TYPE "KP8 Driver: Parameters: 1 Button"
   STRUCT
      activate : Bool;   // true = button on, flase = button off
      cOn1 : String[10];   // color when button is in pressed state. valid entries: 'red', 'green', 'blue', 'yellow', 'white', 'off'
      cOn2 : String[10];   // second flash color when button is pressed and flashing is enabled. valid entries: 'red', 'green', 'blue', 'yellow', 'white', 'off'
      cOff : String[10];   // color when button is in un-pressed state. valid entries: 'red', 'green', 'blue', 'yellow', 'white', 'off'
      flash : Bool;   // false = color 1, true = color 2. set to clock bit to flash at that rate
      group : Int;   // 0 disables. buttons in groups have a mutually exclusive 'on' state.
      mode : Bool;   // true = maintained, fales = momentary
   END_STRUCT;
END_TYPE

TYPE "Selectable Wips"
   STRUCT
      count : Int;
      wips : Array[0.."wipCount"] of DInt;
   END_STRUCT;
END_TYPE

TYPE "Recipe: PN Text Library"
VERSION : 0.1
   STRUCT
      pnText : Array[0.."pnLibCount"] of WString["sStringLen"];
   END_STRUCT;
END_TYPE

TYPE "Selected Wips"
   STRUCT
      count : Int;
      wips : Array[0.."wipCount"] of DInt;
   END_STRUCT;
END_TYPE

TYPE "Selected Buttons"
   STRUCT
      btns : Array[0.."btnCount"] of Bool;
      count : Int;
   END_STRUCT;
END_TYPE

TYPE "KP8 Driver: Button States"
   STRUCT
      btn : Array[0..7] of Bool;
   END_STRUCT;
END_TYPE

TYPE "KP8 Driver: Parameters: 8 Buttons"
   STRUCT
      btn : Array[0..7] of "KP8 Driver: Parameters: 1 Button";
   END_STRUCT;
END_TYPE

TYPE "KP8 Driver: Feedback Data"
   STRUCT
      acutal : "KP8 Driver: Button States";
      falling : "KP8 Driver: Button States";
      rising : "KP8 Driver: Button States";
   END_STRUCT;
END_TYPE

TYPE "Setting Meta Data"
   STRUCT
      selectable_stations : "Selectable Stations";
      selectable_wips : "Selectable Wips";
      selected_btns : "Selected Buttons";
      selected_stations : "Selected Stations";
      selected_wips : "Selected Wips";
      selection_change : "Station Selection Change";
   END_STRUCT;
END_TYPE

TYPE "Nav Bar Data"
   STRUCT
      hmi : "Nav Bar Data: HMI";
      plc : "Nav Bar Data: PLC";
   END_STRUCT;
END_TYPE

TYPE "Intersecting WIPs Arrays"
   STRUCT
      count : Int;
      WIPS_intersection : Array[0.."wipCount"] of DInt;
   END_STRUCT;
END_TYPE

TYPE "Initialize Excel Data: States"
   STRUCT
      active_wip_to_hmi_station_list : Bool;
      active_wip_to_master_station_list : Bool;
      pn_code_to_kp8_station : Bool;
      pn_code_to_saved_wips : Bool;
      wip_code_to_saved_wips : Bool;
   END_STRUCT;
END_TYPE

DATA_BLOCK "EMP IDB"   // DB1
{ S7_Optimized_Access := 'TRUE' }
VERSION : 0.1
// stored: InstanceOfName EMP
"EMP"
BEGIN
   "inst HMI Station"."inst HMI Station: Wip Selection".rowIndicies[1] := 1;
   "inst HMI Station"."inst HMI Station: Wip Selection".rowIndicies[2] := 2;
   "inst HMI Station"."inst HMI Station: Wip Selection".rowIndicies[3] := 3;
   "inst HMI Station"."inst HMI Station: Wip Selection".rowIndicies[4] := 4;
   "inst HMI Station"."inst HMI Station: Wip Selection".rowIndicies[5] := 5;
END_DATA_BLOCK

DATA_BLOCK "Debug"   // DB7
{ S7_Optimized_Access := 'TRUE' }
VERSION : 0.1
   VAR
      nullCheck : Array[0.."wipCount"] of DInt;
   END_VAR
BEGIN
END_DATA_BLOCK

// folder: From Excel

DATA_BLOCK "From Excel: Codes"   // DB12
{ S7_Optimized_Access := 'TRUE' }
VERSION : 0.1
BEGIN
   kp8Stns[0].pnCode[0] := 0;
   kp8Stns[0].pnCode[1] := 0;
   kp8Stns[0].pnCode[2] := 0;
   kp8Stns[0].pnCode[3] := 172000;
   kp8Stns[0].pnCode[4] := 0;
   kp8Stns[0].pnCode[5] := 0;
   kp8Stns[0].pnCode[6] := 0;
   kp8Stns[0].pnCode[7] := 168000;
   kp8Stns[1].pnCode[0] := 0;
   kp8Stns[1].pnCode[1] := 0;
   kp8Stns[1].pnCode[2] := 183000;
   kp8Stns[1].pnCode[3] := 209000;
   kp8Stns[1].pnCode[4] := 0;
   kp8Stns[1].pnCode[5] := 0;
   kp8Stns[1].pnCode[6] := 180000;
   kp8Stns[1].pnCode[7] := 166000;
   kp8Stns[2].pnCode[0] := 0;
   kp8Stns[2].pnCode[1] := 182000;
   kp8Stns[2].pnCode[2] := 181000;
   kp8Stns[2].pnCode[3] := 215000;
   kp8Stns[2].pnCode[4] := 0;
   kp8Stns[2].pnCode[5] := 184000;
   kp8Stns[2].pnCode[6] := 216000;
   kp8Stns[2].pnCode[7] := 214000;
   kp8Stns[3].pnCode[0] := 0;
   kp8Stns[3].pnCode[1] := 192000;
   kp8Stns[3].pnCode[2] := 191000;
   kp8Stns[3].pnCode[3] := 188000;
   kp8Stns[3].pnCode[4] := 0;
   kp8Stns[3].pnCode[5] := 190000;
   kp8Stns[3].pnCode[6] := 187000;
   kp8Stns[3].pnCode[7] := 189000;
   kp8Stns[4].pnCode[0] := 0;
   kp8Stns[4].pnCode[1] := 0;
   kp8Stns[4].pnCode[2] := 0;
   kp8Stns[4].pnCode[3] := 0;
   kp8Stns[4].pnCode[4] := 0;
   kp8Stns[4].pnCode[5] := 0;
   kp8Stns[4].pnCode[6] := 0;
   kp8Stns[4].pnCode[7] := 194000;
   kp8Stns[5].pnCode[0] := 0;
   kp8Stns[5].pnCode[1] := 193000;
   kp8Stns[5].pnCode[2] := 195000;
   kp8Stns[5].pnCode[3] := 176000;
   kp8Stns[5].pnCode[4] := 0;
   kp8Stns[5].pnCode[5] := 196000;
   kp8Stns[5].pnCode[6] := 177000;
   kp8Stns[5].pnCode[7] := 175000;
   kp8Stns[6].pnCode[0] := 0;
   kp8Stns[6].pnCode[1] := 208000;
   kp8Stns[6].pnCode[2] := 207000;
   kp8Stns[6].pnCode[3] := 210000;
   kp8Stns[6].pnCode[4] := 0;
   kp8Stns[6].pnCode[5] := 211000;
   kp8Stns[6].pnCode[6] := 206000;
   kp8Stns[6].pnCode[7] := 205000;
   kp8Stns[7].pnCode[0] := 0;
   kp8Stns[7].pnCode[1] := 0;
   kp8Stns[7].pnCode[2] := 0;
   kp8Stns[7].pnCode[3] := 174000;
   kp8Stns[7].pnCode[4] := 0;
   kp8Stns[7].pnCode[5] := 0;
   kp8Stns[7].pnCode[6] := 167000;
   kp8Stns[7].pnCode[7] := 169000;
   kp8Stns[8].pnCode[0] := 0;
   kp8Stns[8].pnCode[1] := 0;
   kp8Stns[8].pnCode[2] := 0;
   kp8Stns[8].pnCode[3] := 204000;
   kp8Stns[8].pnCode[4] := 0;
   kp8Stns[8].pnCode[5] := 0;
   kp8Stns[8].pnCode[6] := 173000;
   kp8Stns[8].pnCode[7] := 186000;
   kp8Stns[9].pnCode[0] := 0;
   kp8Stns[9].pnCode[1] := 0;
   kp8Stns[9].pnCode[2] := 0;
   kp8Stns[9].pnCode[3] := 213000;
   kp8Stns[9].pnCode[4] := 0;
   kp8Stns[9].pnCode[5] := 0;
   kp8Stns[9].pnCode[6] := 0;
   kp8Stns[9].pnCode[7] := 212000;
   kp8Stns[10].pnCode[0] := 0;
   kp8Stns[10].pnCode[1] := 0;
   kp8Stns[10].pnCode[2] := 0;
   kp8Stns[10].pnCode[3] := 170000;
   kp8Stns[10].pnCode[4] := 0;
   kp8Stns[10].pnCode[5] := 0;
   kp8Stns[10].pnCode[6] := 242000;
   kp8Stns[10].pnCode[7] := 171000;
   kp8Stns[11].pnCode[0] := 0;
   kp8Stns[11].pnCode[1] := 0;
   kp8Stns[11].pnCode[2] := 0;
   kp8Stns[11].pnCode[3] := 77000;
   kp8Stns[11].pnCode[4] := 0;
   kp8Stns[11].pnCode[5] := 0;
   kp8Stns[11].pnCode[6] := 65000;
   kp8Stns[11].pnCode[7] := 20000;
   kp8Stns[12].pnCode[0] := 0;
   kp8Stns[12].pnCode[1] := 80000;
   kp8Stns[12].pnCode[2] := 86000;
   kp8Stns[12].pnCode[3] := 59000;
   kp8Stns[12].pnCode[4] := 0;
   kp8Stns[12].pnCode[5] := 79000;
   kp8Stns[12].pnCode[6] := 55000;
   kp8Stns[12].pnCode[7] := 54000;
   kp8Stns[13].pnCode[0] := 0;
   kp8Stns[13].pnCode[1] := 0;
   kp8Stns[13].pnCode[2] := 69000;
   kp8Stns[13].pnCode[3] := 89000;
   kp8Stns[13].pnCode[4] := 0;
   kp8Stns[13].pnCode[5] := 0;
   kp8Stns[13].pnCode[6] := 90000;
   kp8Stns[13].pnCode[7] := 88000;
   kp8Stns[14].pnCode[0] := 0;
   kp8Stns[14].pnCode[1] := 0;
   kp8Stns[14].pnCode[2] := 64000;
   kp8Stns[14].pnCode[3] := 87000;
   kp8Stns[14].pnCode[4] := 0;
   kp8Stns[14].pnCode[5] := 63000;
   kp8Stns[14].pnCode[6] := 82000;
   kp8Stns[14].pnCode[7] := 62000;
   kp8Stns[15].pnCode[0] := 0;
   kp8Stns[15].pnCode[1] := 49000;
   kp8Stns[15].pnCode[2] := 76000;
   kp8Stns[15].pnCode[3] := 28000;
   kp8Stns[15].pnCode[4] := 0;
   kp8Stns[15].pnCode[5] := 81000;
   kp8Stns[15].pnCode[6] := 68000;
   kp8Stns[15].pnCode[7] := 74000;
   kp8Stns[16].pnCode[0] := 0;
   kp8Stns[16].pnCode[1] := 0;
   kp8Stns[16].pnCode[2] := 0;
   kp8Stns[16].pnCode[3] := 91000;
   kp8Stns[16].pnCode[4] := 0;
   kp8Stns[16].pnCode[5] := 0;
   kp8Stns[16].pnCode[6] := 93000;
   kp8Stns[16].pnCode[7] := 94067;
   kp8Stns[17].pnCode[0] := 0;
   kp8Stns[17].pnCode[1] := 0;
   kp8Stns[17].pnCode[2] := 83000;
   kp8Stns[17].pnCode[3] := 34000;
   kp8Stns[17].pnCode[4] := 0;
   kp8Stns[17].pnCode[5] := 0;
   kp8Stns[17].pnCode[6] := 75000;
   kp8Stns[17].pnCode[7] := 29000;
   kp8Stns[18].pnCode[0] := 0;
   kp8Stns[18].pnCode[1] := 0;
   kp8Stns[18].pnCode[2] := 0;
   kp8Stns[18].pnCode[3] := 92066;
   kp8Stns[18].pnCode[4] := 0;
   kp8Stns[18].pnCode[5] := 0;
   kp8Stns[18].pnCode[6] := 96026;
   kp8Stns[18].pnCode[7] := 95000;
   kp8Stns[19].pnCode[0] := 0;
   kp8Stns[19].pnCode[1] := 78000;
   kp8Stns[19].pnCode[2] := 85000;
   kp8Stns[19].pnCode[3] := 21000;
   kp8Stns[19].pnCode[4] := 0;
   kp8Stns[19].pnCode[5] := 97000;
   kp8Stns[19].pnCode[6] := 60000;
   kp8Stns[19].pnCode[7] := 48000;
   kp8Stns[20].pnCode[0] := 0;
   kp8Stns[20].pnCode[1] := 0;
   kp8Stns[20].pnCode[2] := 0;
   kp8Stns[20].pnCode[3] := 0;
   kp8Stns[20].pnCode[4] := 0;
   kp8Stns[20].pnCode[5] := 0;
   kp8Stns[20].pnCode[6] := 0;
   kp8Stns[20].pnCode[7] := 244000;
   kp8Stns[21].pnCode[0] := 0;
   kp8Stns[21].pnCode[1] := 0;
   kp8Stns[21].pnCode[2] := 0;
   kp8Stns[21].pnCode[3] := 245000;
   kp8Stns[21].pnCode[4] := 0;
   kp8Stns[21].pnCode[5] := 0;
   kp8Stns[21].pnCode[6] := 0;
   kp8Stns[21].pnCode[7] := 11000;
   kp8Stns[22].pnCode[0] := 0;
   kp8Stns[22].pnCode[1] := 0;
   kp8Stns[22].pnCode[2] := 0;
   kp8Stns[22].pnCode[3] := 22000;
   kp8Stns[22].pnCode[4] := 0;
   kp8Stns[22].pnCode[5] := 0;
   kp8Stns[22].pnCode[6] := 46000;
   kp8Stns[22].pnCode[7] := 61000;
   kp8Stns[23].pnCode[0] := 0;
   kp8Stns[23].pnCode[1] := 0;
   kp8Stns[23].pnCode[2] := 0;
   kp8Stns[23].pnCode[3] := 0;
   kp8Stns[23].pnCode[4] := 0;
   kp8Stns[23].pnCode[5] := 0;
   kp8Stns[23].pnCode[6] := 0;
   kp8Stns[23].pnCode[7] := 12000;
   kp8Stns[24].pnCode[0] := 0;
   kp8Stns[24].pnCode[1] := 0;
   kp8Stns[24].pnCode[2] := 0;
   kp8Stns[24].pnCode[3] := 0;
   kp8Stns[24].pnCode[4] := 0;
   kp8Stns[24].pnCode[5] := 0;
   kp8Stns[24].pnCode[6] := 0;
   kp8Stns[24].pnCode[7] := 27000;
   kp8Stns[25].pnCode[0] := 0;
   kp8Stns[25].pnCode[1] := 0;
   kp8Stns[25].pnCode[2] := 0;
   kp8Stns[25].pnCode[3] := 0;
   kp8Stns[25].pnCode[4] := 0;
   kp8Stns[25].pnCode[5] := 0;
   kp8Stns[25].pnCode[6] := 0;
   kp8Stns[25].pnCode[7] := 56000;
   hmiStns[0].wip[0].wipCode := 6027;
   hmiStns[0].wip[0].pnCode[0] := 0;
   hmiStns[0].wip[0].pnCode[1] := 243000;
   hmiStns[0].wip[0].pnCode[2] := 19000;
   hmiStns[0].wip[0].pnCode[3] := 0;
   hmiStns[0].wip[0].pnCode[4] := 0;
   hmiStns[0].wip[0].pnCode[5] := 0;
   hmiStns[0].wip[0].pnCode[6] := 25000;
   hmiStns[0].wip[0].pnCode[7] := 18000;
   hmiStns[0].wip[1].wipCode := 9007;
   hmiStns[0].wip[1].pnCode[0] := 0;
   hmiStns[0].wip[1].pnCode[1] := 243000;
   hmiStns[0].wip[1].pnCode[2] := 37000;
   hmiStns[0].wip[1].pnCode[3] := 0;
   hmiStns[0].wip[1].pnCode[4] := 0;
   hmiStns[0].wip[1].pnCode[5] := 0;
   hmiStns[0].wip[1].pnCode[6] := 35000;
   hmiStns[0].wip[1].pnCode[7] := 36000;
   hmiStns[0].wip[2].wipCode := 10030;
   hmiStns[0].wip[2].pnCode[0] := 0;
   hmiStns[0].wip[2].pnCode[1] := 243000;
   hmiStns[0].wip[2].pnCode[2] := 40000;
   hmiStns[0].wip[2].pnCode[3] := 0;
   hmiStns[0].wip[2].pnCode[4] := 0;
   hmiStns[0].wip[2].pnCode[5] := 0;
   hmiStns[0].wip[2].pnCode[6] := 38000;
   hmiStns[0].wip[2].pnCode[7] := 39000;
   hmiStns[0].wip[3].wipCode := 11056;
   hmiStns[0].wip[3].pnCode[0] := 0;
   hmiStns[0].wip[3].pnCode[1] := 243000;
   hmiStns[0].wip[3].pnCode[2] := 47000;
   hmiStns[0].wip[3].pnCode[3] := 13000;
   hmiStns[0].wip[3].pnCode[4] := 0;
   hmiStns[0].wip[3].pnCode[5] := 14000;
   hmiStns[0].wip[3].pnCode[6] := 41000;
   hmiStns[0].wip[3].pnCode[7] := 32000;
   hmiStns[0].wip[4].wipCode := 12008;
   hmiStns[0].wip[4].pnCode[0] := 0;
   hmiStns[0].wip[4].pnCode[1] := 243000;
   hmiStns[0].wip[4].pnCode[2] := 45000;
   hmiStns[0].wip[4].pnCode[3] := 0;
   hmiStns[0].wip[4].pnCode[4] := 0;
   hmiStns[0].wip[4].pnCode[5] := 0;
   hmiStns[0].wip[4].pnCode[6] := 35000;
   hmiStns[0].wip[4].pnCode[7] := 36000;
   hmiStns[0].wip[5].wipCode := 13060;
   hmiStns[0].wip[5].pnCode[0] := 0;
   hmiStns[0].wip[5].pnCode[1] := 243000;
   hmiStns[0].wip[5].pnCode[2] := 37000;
   hmiStns[0].wip[5].pnCode[3] := 0;
   hmiStns[0].wip[5].pnCode[4] := 0;
   hmiStns[0].wip[5].pnCode[5] := 0;
   hmiStns[0].wip[5].pnCode[6] := 42000;
   hmiStns[0].wip[5].pnCode[7] := 36000;
   hmiStns[0].wip[6].wipCode := 14061;
   hmiStns[0].wip[6].pnCode[0] := 0;
   hmiStns[0].wip[6].pnCode[1] := 243000;
   hmiStns[0].wip[6].pnCode[2] := 45000;
   hmiStns[0].wip[6].pnCode[3] := 0;
   hmiStns[0].wip[6].pnCode[4] := 0;
   hmiStns[0].wip[6].pnCode[5] := 0;
   hmiStns[0].wip[6].pnCode[6] := 42000;
   hmiStns[0].wip[6].pnCode[7] := 36000;
   hmiStns[0].wip[7].wipCode := 15030;
   hmiStns[0].wip[7].pnCode[0] := 0;
   hmiStns[0].wip[7].pnCode[1] := 243000;
   hmiStns[0].wip[7].pnCode[2] := 43000;
   hmiStns[0].wip[7].pnCode[3] := 0;
   hmiStns[0].wip[7].pnCode[4] := 0;
   hmiStns[0].wip[7].pnCode[5] := 0;
   hmiStns[0].wip[7].pnCode[6] := 38000;
   hmiStns[0].wip[7].pnCode[7] := 44000;
   hmiStns[0].wip[8].wipCode := 16024;
   hmiStns[0].wip[8].pnCode[0] := 0;
   hmiStns[0].wip[8].pnCode[1] := 243000;
   hmiStns[0].wip[8].pnCode[2] := 51000;
   hmiStns[0].wip[8].pnCode[3] := 0;
   hmiStns[0].wip[8].pnCode[4] := 0;
   hmiStns[0].wip[8].pnCode[5] := 0;
   hmiStns[0].wip[8].pnCode[6] := 25000;
   hmiStns[0].wip[8].pnCode[7] := 18000;
   hmiStns[0].wip[9].wipCode := 17009;
   hmiStns[0].wip[9].pnCode[0] := 0;
   hmiStns[0].wip[9].pnCode[1] := 243000;
   hmiStns[0].wip[9].pnCode[2] := 52000;
   hmiStns[0].wip[9].pnCode[3] := 0;
   hmiStns[0].wip[9].pnCode[4] := 0;
   hmiStns[0].wip[9].pnCode[5] := 0;
   hmiStns[0].wip[9].pnCode[6] := 31000;
   hmiStns[0].wip[9].pnCode[7] := 73000;
   hmiStns[0].wip[10].wipCode := 19031;
   hmiStns[0].wip[10].pnCode[0] := 0;
   hmiStns[0].wip[10].pnCode[1] := 243000;
   hmiStns[0].wip[10].pnCode[2] := 53000;
   hmiStns[0].wip[10].pnCode[3] := 0;
   hmiStns[0].wip[10].pnCode[4] := 0;
   hmiStns[0].wip[10].pnCode[5] := 0;
   hmiStns[0].wip[10].pnCode[6] := 31000;
   hmiStns[0].wip[10].pnCode[7] := 71000;
   hmiStns[0].wip[11].wipCode := 21028;
   hmiStns[0].wip[11].pnCode[0] := 0;
   hmiStns[0].wip[11].pnCode[1] := 243000;
   hmiStns[0].wip[11].pnCode[2] := 57000;
   hmiStns[0].wip[11].pnCode[3] := 0;
   hmiStns[0].wip[11].pnCode[4] := 0;
   hmiStns[0].wip[11].pnCode[5] := 0;
   hmiStns[0].wip[11].pnCode[6] := 25000;
   hmiStns[0].wip[11].pnCode[7] := 18000;
   hmiStns[0].wip[12].wipCode := 22008;
   hmiStns[0].wip[12].pnCode[0] := 0;
   hmiStns[0].wip[12].pnCode[1] := 243000;
   hmiStns[0].wip[12].pnCode[2] := 84000;
   hmiStns[0].wip[12].pnCode[3] := 0;
   hmiStns[0].wip[12].pnCode[4] := 0;
   hmiStns[0].wip[12].pnCode[5] := 0;
   hmiStns[0].wip[12].pnCode[6] := 31000;
   hmiStns[0].wip[12].pnCode[7] := 71000;
   hmiStns[0].wip[13].wipCode := 24029;
   hmiStns[0].wip[13].pnCode[0] := 0;
   hmiStns[0].wip[13].pnCode[1] := 243000;
   hmiStns[0].wip[13].pnCode[2] := 98000;
   hmiStns[0].wip[13].pnCode[3] := 0;
   hmiStns[0].wip[13].pnCode[4] := 0;
   hmiStns[0].wip[13].pnCode[5] := 0;
   hmiStns[0].wip[13].pnCode[6] := 38000;
   hmiStns[0].wip[13].pnCode[7] := 44000;
   hmiStns[0].wip[14].wipCode := 25025;
   hmiStns[0].wip[14].pnCode[0] := 0;
   hmiStns[0].wip[14].pnCode[1] := 243000;
   hmiStns[0].wip[14].pnCode[2] := 99000;
   hmiStns[0].wip[14].pnCode[3] := 0;
   hmiStns[0].wip[14].pnCode[4] := 0;
   hmiStns[0].wip[14].pnCode[5] := 0;
   hmiStns[0].wip[14].pnCode[6] := 42000;
   hmiStns[0].wip[14].pnCode[7] := 36000;
   hmiStns[0].wip[15].wipCode := 26026;
   hmiStns[0].wip[15].pnCode[0] := 0;
   hmiStns[0].wip[15].pnCode[1] := 243000;
   hmiStns[0].wip[15].pnCode[2] := 99000;
   hmiStns[0].wip[15].pnCode[3] := 0;
   hmiStns[0].wip[15].pnCode[4] := 0;
   hmiStns[0].wip[15].pnCode[5] := 0;
   hmiStns[0].wip[15].pnCode[6] := 35000;
   hmiStns[0].wip[15].pnCode[7] := 36000;
   hmiStns[0].wip[16].wipCode := 69063;
   hmiStns[0].wip[16].pnCode[0] := 0;
   hmiStns[0].wip[16].pnCode[1] := 243000;
   hmiStns[0].wip[16].pnCode[2] := 217000;
   hmiStns[0].wip[16].pnCode[3] := 0;
   hmiStns[0].wip[16].pnCode[4] := 0;
   hmiStns[0].wip[16].pnCode[5] := 0;
   hmiStns[0].wip[16].pnCode[6] := 218000;
   hmiStns[0].wip[16].pnCode[7] := 223000;
   hmiStns[0].wip[17].wipCode := 71000;
   hmiStns[0].wip[17].pnCode[0] := 0;
   hmiStns[0].wip[17].pnCode[1] := 243000;
   hmiStns[0].wip[17].pnCode[2] := 197000;
   hmiStns[0].wip[17].pnCode[3] := 0;
   hmiStns[0].wip[17].pnCode[4] := 0;
   hmiStns[0].wip[17].pnCode[5] := 0;
   hmiStns[0].wip[17].pnCode[6] := 219000;
   hmiStns[0].wip[17].pnCode[7] := 222000;
   hmiStns[0].wip[18].wipCode := 72023;
   hmiStns[0].wip[18].pnCode[0] := 0;
   hmiStns[0].wip[18].pnCode[1] := 243000;
   hmiStns[0].wip[18].pnCode[2] := 198000;
   hmiStns[0].wip[18].pnCode[3] := 0;
   hmiStns[0].wip[18].pnCode[4] := 0;
   hmiStns[0].wip[18].pnCode[5] := 0;
   hmiStns[0].wip[18].pnCode[6] := 218000;
   hmiStns[0].wip[18].pnCode[7] := 223000;
   hmiStns[0].wip[19].wipCode := 73064;
   hmiStns[0].wip[19].pnCode[0] := 0;
   hmiStns[0].wip[19].pnCode[1] := 243000;
   hmiStns[0].wip[19].pnCode[2] := 224000;
   hmiStns[0].wip[19].pnCode[3] := 0;
   hmiStns[0].wip[19].pnCode[4] := 0;
   hmiStns[0].wip[19].pnCode[5] := 0;
   hmiStns[0].wip[19].pnCode[6] := 225000;
   hmiStns[0].wip[19].pnCode[7] := 226000;
   hmiStns[0].wip[20].wipCode := 5009;
   hmiStns[0].wip[20].pnCode[0] := 0;
   hmiStns[0].wip[20].pnCode[1] := 243000;
   hmiStns[0].wip[20].pnCode[2] := 17000;
   hmiStns[0].wip[20].pnCode[3] := 0;
   hmiStns[0].wip[20].pnCode[4] := 0;
   hmiStns[0].wip[20].pnCode[5] := 0;
   hmiStns[0].wip[20].pnCode[6] := 24000;
   hmiStns[0].wip[20].pnCode[7] := 16000;
   hmiStns[0].wip[21].wipCode := 7031;
   hmiStns[0].wip[21].pnCode[0] := 0;
   hmiStns[0].wip[21].pnCode[1] := 243000;
   hmiStns[0].wip[21].pnCode[2] := 0;
   hmiStns[0].wip[21].pnCode[3] := 31000;
   hmiStns[0].wip[21].pnCode[4] := 0;
   hmiStns[0].wip[21].pnCode[5] := 0;
   hmiStns[0].wip[21].pnCode[6] := 50000;
   hmiStns[0].wip[21].pnCode[7] := 30000;
   hmiStns[0].wip[22].wipCode := 74011;
   hmiStns[0].wip[22].pnCode[0] := 0;
   hmiStns[0].wip[22].pnCode[1] := 243000;
   hmiStns[0].wip[22].pnCode[2] := 0;
   hmiStns[0].wip[22].pnCode[3] := 219000;
   hmiStns[0].wip[22].pnCode[4] := 0;
   hmiStns[0].wip[22].pnCode[5] := 0;
   hmiStns[0].wip[22].pnCode[6] := 221000;
   hmiStns[0].wip[22].pnCode[7] := 222000;
   hmiStns[0].wip[23].wipCode := 70010;
   hmiStns[0].wip[23].pnCode[0] := 0;
   hmiStns[0].wip[23].pnCode[1] := 243000;
   hmiStns[0].wip[23].pnCode[2] := 220000;
   hmiStns[0].wip[23].pnCode[3] := 0;
   hmiStns[0].wip[23].pnCode[4] := 0;
   hmiStns[0].wip[23].pnCode[5] := 0;
   hmiStns[0].wip[23].pnCode[6] := 219000;
   hmiStns[0].wip[23].pnCode[7] := 222000;
   hmiStns[0].wip[24].wipCode := -1;
   hmiStns[0].wip[24].pnCode[0] := 0;
   hmiStns[0].wip[24].pnCode[1] := 0;
   hmiStns[0].wip[24].pnCode[2] := 0;
   hmiStns[0].wip[24].pnCode[3] := 0;
   hmiStns[0].wip[24].pnCode[4] := 0;
   hmiStns[0].wip[24].pnCode[5] := 0;
   hmiStns[0].wip[24].pnCode[6] := 0;
   hmiStns[0].wip[24].pnCode[7] := 0;
   hmiStns[0].wip[25].wipCode := -1;
   hmiStns[0].wip[25].pnCode[0] := 0;
   hmiStns[0].wip[25].pnCode[1] := 0;
   hmiStns[0].wip[25].pnCode[2] := 0;
   hmiStns[0].wip[25].pnCode[3] := 0;
   hmiStns[0].wip[25].pnCode[4] := 0;
   hmiStns[0].wip[25].pnCode[5] := 0;
   hmiStns[0].wip[25].pnCode[6] := 0;
   hmiStns[0].wip[25].pnCode[7] := 0;
   hmiStns[0].wip[26].wipCode := -1;
   hmiStns[0].wip[26].pnCode[0] := 0;
   hmiStns[0].wip[26].pnCode[1] := 0;
   hmiStns[0].wip[26].pnCode[2] := 0;
   hmiStns[0].wip[26].pnCode[3] := 0;
   hmiStns[0].wip[26].pnCode[4] := 0;
   hmiStns[0].wip[26].pnCode[5] := 0;
   hmiStns[0].wip[26].pnCode[6] := 0;
   hmiStns[0].wip[26].pnCode[7] := 0;
   hmiStns[0].wip[27].wipCode := -1;
   hmiStns[0].wip[27].pnCode[0] := 0;
   hmiStns[0].wip[27].pnCode[1] := 0;
   hmiStns[0].wip[27].pnCode[2] := 0;
   hmiStns[0].wip[27].pnCode[3] := 0;
   hmiStns[0].wip[27].pnCode[4] := 0;
   hmiStns[0].wip[27].pnCode[5] := 0;
   hmiStns[0].wip[27].pnCode[6] := 0;
   hmiStns[0].wip[27].pnCode[7] := 0;
   hmiStns[0].wip[28].wipCode := -1;
   hmiStns[0].wip[28].pnCode[0] := 0;
   hmiStns[0].wip[28].pnCode[1] := 0;
   hmiStns[0].wip[28].pnCode[2] := 0;
   hmiStns[0].wip[28].pnCode[3] := 0;
   hmiStns[0].wip[28].pnCode[4] := 0;
   hmiStns[0].wip[28].pnCode[5] := 0;
   hmiStns[0].wip[28].pnCode[6] := 0;
   hmiStns[0].wip[28].pnCode[7] := 0;
   hmiStns[0].wip[29].wipCode := -1;
   hmiStns[0].wip[29].pnCode[0] := 0;
   hmiStns[0].wip[29].pnCode[1] := 0;
   hmiStns[0].wip[29].pnCode[2] := 0;
   hmiStns[0].wip[29].pnCode[3] := 0;
   hmiStns[0].wip[29].pnCode[4] := 0;
   hmiStns[0].wip[29].pnCode[5] := 0;
   hmiStns[0].wip[29].pnCode[6] := 0;
   hmiStns[0].wip[29].pnCode[7] := 0;
   hmiStns[0].wip[30].wipCode := -1;
   hmiStns[0].wip[30].pnCode[0] := 0;
   hmiStns[0].wip[30].pnCode[1] := 0;
   hmiStns[0].wip[30].pnCode[2] := 0;
   hmiStns[0].wip[30].pnCode[3] := 0;
   hmiStns[0].wip[30].pnCode[4] := 0;
   hmiStns[0].wip[30].pnCode[5] := 0;
   hmiStns[0].wip[30].pnCode[6] := 0;
   hmiStns[0].wip[30].pnCode[7] := 0;
   hmiStns[0].wip[31].wipCode := -1;
   hmiStns[0].wip[31].pnCode[0] := 0;
   hmiStns[0].wip[31].pnCode[1] := 0;
   hmiStns[0].wip[31].pnCode[2] := 0;
   hmiStns[0].wip[31].pnCode[3] := 0;
   hmiStns[0].wip[31].pnCode[4] := 0;
   hmiStns[0].wip[31].pnCode[5] := 0;
   hmiStns[0].wip[31].pnCode[6] := 0;
   hmiStns[0].wip[31].pnCode[7] := 0;
   hmiStns[0].wip[32].wipCode := -1;
   hmiStns[0].wip[32].pnCode[0] := 0;
   hmiStns[0].wip[32].pnCode[1] := 0;
   hmiStns[0].wip[32].pnCode[2] := 0;
   hmiStns[0].wip[32].pnCode[3] := 0;
   hmiStns[0].wip[32].pnCode[4] := 0;
   hmiStns[0].wip[32].pnCode[5] := 0;
   hmiStns[0].wip[32].pnCode[6] := 0;
   hmiStns[0].wip[32].pnCode[7] := 0;
   hmiStns[0].wip[33].wipCode := -1;
   hmiStns[0].wip[33].pnCode[0] := 0;
   hmiStns[0].wip[33].pnCode[1] := 0;
   hmiStns[0].wip[33].pnCode[2] := 0;
   hmiStns[0].wip[33].pnCode[3] := 0;
   hmiStns[0].wip[33].pnCode[4] := 0;
   hmiStns[0].wip[33].pnCode[5] := 0;
   hmiStns[0].wip[33].pnCode[6] := 0;
   hmiStns[0].wip[33].pnCode[7] := 0;
   hmiStns[0].wip[34].wipCode := -1;
   hmiStns[0].wip[34].pnCode[0] := 0;
   hmiStns[0].wip[34].pnCode[1] := 0;
   hmiStns[0].wip[34].pnCode[2] := 0;
   hmiStns[0].wip[34].pnCode[3] := 0;
   hmiStns[0].wip[34].pnCode[4] := 0;
   hmiStns[0].wip[34].pnCode[5] := 0;
   hmiStns[0].wip[34].pnCode[6] := 0;
   hmiStns[0].wip[34].pnCode[7] := 0;
   hmiStns[0].wip[35].wipCode := -1;
   hmiStns[0].wip[35].pnCode[0] := 0;
   hmiStns[0].wip[35].pnCode[1] := 0;
   hmiStns[0].wip[35].pnCode[2] := 0;
   hmiStns[0].wip[35].pnCode[3] := 0;
   hmiStns[0].wip[35].pnCode[4] := 0;
   hmiStns[0].wip[35].pnCode[5] := 0;
   hmiStns[0].wip[35].pnCode[6] := 0;
   hmiStns[0].wip[35].pnCode[7] := 0;
   hmiStns[0].wip[36].wipCode := -1;
   hmiStns[0].wip[36].pnCode[0] := 0;
   hmiStns[0].wip[36].pnCode[1] := 0;
   hmiStns[0].wip[36].pnCode[2] := 0;
   hmiStns[0].wip[36].pnCode[3] := 0;
   hmiStns[0].wip[36].pnCode[4] := 0;
   hmiStns[0].wip[36].pnCode[5] := 0;
   hmiStns[0].wip[36].pnCode[6] := 0;
   hmiStns[0].wip[36].pnCode[7] := 0;
   hmiStns[0].wip[37].wipCode := -1;
   hmiStns[0].wip[37].pnCode[0] := 0;
   hmiStns[0].wip[37].pnCode[1] := 0;
   hmiStns[0].wip[37].pnCode[2] := 0;
   hmiStns[0].wip[37].pnCode[3] := 0;
   hmiStns[0].wip[37].pnCode[4] := 0;
   hmiStns[0].wip[37].pnCode[5] := 0;
   hmiStns[0].wip[37].pnCode[6] := 0;
   hmiStns[0].wip[37].pnCode[7] := 0;
   hmiStns[0].wip[38].wipCode := -1;
   hmiStns[0].wip[38].pnCode[0] := 0;
   hmiStns[0].wip[38].pnCode[1] := 0;
   hmiStns[0].wip[38].pnCode[2] := 0;
   hmiStns[0].wip[38].pnCode[3] := 0;
   hmiStns[0].wip[38].pnCode[4] := 0;
   hmiStns[0].wip[38].pnCode[5] := 0;
   hmiStns[0].wip[38].pnCode[6] := 0;
   hmiStns[0].wip[38].pnCode[7] := 0;
   hmiStns[0].wip[39].wipCode := -1;
   hmiStns[0].wip[39].pnCode[0] := 0;
   hmiStns[0].wip[39].pnCode[1] := 0;
   hmiStns[0].wip[39].pnCode[2] := 0;
   hmiStns[0].wip[39].pnCode[3] := 0;
   hmiStns[0].wip[39].pnCode[4] := 0;
   hmiStns[0].wip[39].pnCode[5] := 0;
   hmiStns[0].wip[39].pnCode[6] := 0;
   hmiStns[0].wip[39].pnCode[7] := 0;
   hmiStns[0].wip[40].wipCode := -1;
   hmiStns[0].wip[40].pnCode[0] := 0;
   hmiStns[0].wip[40].pnCode[1] := 0;
   hmiStns[0].wip[40].pnCode[2] := 0;
   hmiStns[0].wip[40].pnCode[3] := 0;
   hmiStns[0].wip[40].pnCode[4] := 0;
   hmiStns[0].wip[40].pnCode[5] := 0;
   hmiStns[0].wip[40].pnCode[6] := 0;
   hmiStns[0].wip[40].pnCode[7] := 0;
   hmiStns[0].wip[41].wipCode := -1;
   hmiStns[0].wip[41].pnCode[0] := 0;
   hmiStns[0].wip[41].pnCode[1] := 0;
   hmiStns[0].wip[41].pnCode[2] := 0;
   hmiStns[0].wip[41].pnCode[3] := 0;
   hmiStns[0].wip[41].pnCode[4] := 0;
   hmiStns[0].wip[41].pnCode[5] := 0;
   hmiStns[0].wip[41].pnCode[6] := 0;
   hmiStns[0].wip[41].pnCode[7] := 0;
   hmiStns[0].wip[42].wipCode := -1;
   hmiStns[0].wip[42].pnCode[0] := 0;
   hmiStns[0].wip[42].pnCode[1] := 0;
   hmiStns[0].wip[42].pnCode[2] := 0;
   hmiStns[0].wip[42].pnCode[3] := 0;
   hmiStns[0].wip[42].pnCode[4] := 0;
   hmiStns[0].wip[42].pnCode[5] := 0;
   hmiStns[0].wip[42].pnCode[6] := 0;
   hmiStns[0].wip[42].pnCode[7] := 0;
   hmiStns[0].wip[43].wipCode := -1;
   hmiStns[0].wip[43].pnCode[0] := 0;
   hmiStns[0].wip[43].pnCode[1] := 0;
   hmiStns[0].wip[43].pnCode[2] := 0;
   hmiStns[0].wip[43].pnCode[3] := 0;
   hmiStns[0].wip[43].pnCode[4] := 0;
   hmiStns[0].wip[43].pnCode[5] := 0;
   hmiStns[0].wip[43].pnCode[6] := 0;
   hmiStns[0].wip[43].pnCode[7] := 0;
   hmiStns[0].wip[44].wipCode := -1;
   hmiStns[0].wip[44].pnCode[0] := 0;
   hmiStns[0].wip[44].pnCode[1] := 0;
   hmiStns[0].wip[44].pnCode[2] := 0;
   hmiStns[0].wip[44].pnCode[3] := 0;
   hmiStns[0].wip[44].pnCode[4] := 0;
   hmiStns[0].wip[44].pnCode[5] := 0;
   hmiStns[0].wip[44].pnCode[6] := 0;
   hmiStns[0].wip[44].pnCode[7] := 0;
   hmiStns[0].wip[45].wipCode := -1;
   hmiStns[0].wip[45].pnCode[0] := 0;
   hmiStns[0].wip[45].pnCode[1] := 0;
   hmiStns[0].wip[45].pnCode[2] := 0;
   hmiStns[0].wip[45].pnCode[3] := 0;
   hmiStns[0].wip[45].pnCode[4] := 0;
   hmiStns[0].wip[45].pnCode[5] := 0;
   hmiStns[0].wip[45].pnCode[6] := 0;
   hmiStns[0].wip[45].pnCode[7] := 0;
   hmiStns[0].wip[46].wipCode := -1;
   hmiStns[0].wip[46].pnCode[0] := 0;
   hmiStns[0].wip[46].pnCode[1] := 0;
   hmiStns[0].wip[46].pnCode[2] := 0;
   hmiStns[0].wip[46].pnCode[3] := 0;
   hmiStns[0].wip[46].pnCode[4] := 0;
   hmiStns[0].wip[46].pnCode[5] := 0;
   hmiStns[0].wip[46].pnCode[6] := 0;
   hmiStns[0].wip[46].pnCode[7] := 0;
   hmiStns[0].wip[47].wipCode := -1;
   hmiStns[0].wip[47].pnCode[0] := 0;
   hmiStns[0].wip[47].pnCode[1] := 0;
   hmiStns[0].wip[47].pnCode[2] := 0;
   hmiStns[0].wip[47].pnCode[3] := 0;
   hmiStns[0].wip[47].pnCode[4] := 0;
   hmiStns[0].wip[47].pnCode[5] := 0;
   hmiStns[0].wip[47].pnCode[6] := 0;
   hmiStns[0].wip[47].pnCode[7] := 0;
   hmiStns[0].wip[48].wipCode := -1;
   hmiStns[0].wip[48].pnCode[0] := 0;
   hmiStns[0].wip[48].pnCode[1] := 0;
   hmiStns[0].wip[48].pnCode[2] := 0;
   hmiStns[0].wip[48].pnCode[3] := 0;
   hmiStns[0].wip[48].pnCode[4] := 0;
   hmiStns[0].wip[48].pnCode[5] := 0;
   hmiStns[0].wip[48].pnCode[6] := 0;
   hmiStns[0].wip[48].pnCode[7] := 0;
   hmiStns[0].wip[49].wipCode := -1;
   hmiStns[0].wip[49].pnCode[0] := 0;
   hmiStns[0].wip[49].pnCode[1] := 0;
   hmiStns[0].wip[49].pnCode[2] := 0;
   hmiStns[0].wip[49].pnCode[3] := 0;
   hmiStns[0].wip[49].pnCode[4] := 0;
   hmiStns[0].wip[49].pnCode[5] := 0;
   hmiStns[0].wip[49].pnCode[6] := 0;
   hmiStns[0].wip[49].pnCode[7] := 0;
   hmiStns[1].wip[0].wipCode := 14061;
   hmiStns[1].wip[0].pnCode[0] := 0;
   hmiStns[1].wip[0].pnCode[1] := 243000;
   hmiStns[1].wip[0].pnCode[2] := 45000;
   hmiStns[1].wip[0].pnCode[3] := 0;
   hmiStns[1].wip[0].pnCode[4] := 0;
   hmiStns[1].wip[0].pnCode[5] := 0;
   hmiStns[1].wip[0].pnCode[6] := 42000;
   hmiStns[1].wip[0].pnCode[7] := 36000;
   hmiStns[1].wip[1].wipCode := 25025;
   hmiStns[1].wip[1].pnCode[0] := 0;
   hmiStns[1].wip[1].pnCode[1] := 243000;
   hmiStns[1].wip[1].pnCode[2] := 99000;
   hmiStns[1].wip[1].pnCode[3] := 0;
   hmiStns[1].wip[1].pnCode[4] := 0;
   hmiStns[1].wip[1].pnCode[5] := 0;
   hmiStns[1].wip[1].pnCode[6] := 42000;
   hmiStns[1].wip[1].pnCode[7] := 36000;
   hmiStns[1].wip[2].wipCode := 26026;
   hmiStns[1].wip[2].pnCode[0] := 0;
   hmiStns[1].wip[2].pnCode[1] := 243000;
   hmiStns[1].wip[2].pnCode[2] := 99000;
   hmiStns[1].wip[2].pnCode[3] := 0;
   hmiStns[1].wip[2].pnCode[4] := 0;
   hmiStns[1].wip[2].pnCode[5] := 0;
   hmiStns[1].wip[2].pnCode[6] := 35000;
   hmiStns[1].wip[2].pnCode[7] := 36000;
   hmiStns[1].wip[3].wipCode := 4052;
   hmiStns[1].wip[3].pnCode[0] := 0;
   hmiStns[1].wip[3].pnCode[1] := 243000;
   hmiStns[1].wip[3].pnCode[2] := 14000;
   hmiStns[1].wip[3].pnCode[3] := 0;
   hmiStns[1].wip[3].pnCode[4] := 0;
   hmiStns[1].wip[3].pnCode[5] := 15000;
   hmiStns[1].wip[3].pnCode[6] := 23000;
   hmiStns[1].wip[3].pnCode[7] := 13000;
   hmiStns[1].wip[4].wipCode := 8062;
   hmiStns[1].wip[4].pnCode[0] := 0;
   hmiStns[1].wip[4].pnCode[1] := 243000;
   hmiStns[1].wip[4].pnCode[2] := 14000;
   hmiStns[1].wip[4].pnCode[3] := 13000;
   hmiStns[1].wip[4].pnCode[4] := 0;
   hmiStns[1].wip[4].pnCode[5] := 47000;
   hmiStns[1].wip[4].pnCode[6] := 33000;
   hmiStns[1].wip[4].pnCode[7] := 32000;
   hmiStns[1].wip[5].wipCode := 18053;
   hmiStns[1].wip[5].pnCode[0] := 0;
   hmiStns[1].wip[5].pnCode[1] := 243000;
   hmiStns[1].wip[5].pnCode[2] := 14000;
   hmiStns[1].wip[5].pnCode[3] := 0;
   hmiStns[1].wip[5].pnCode[4] := 0;
   hmiStns[1].wip[5].pnCode[5] := 15000;
   hmiStns[1].wip[5].pnCode[6] := 33000;
   hmiStns[1].wip[5].pnCode[7] := 13000;
   hmiStns[1].wip[6].wipCode := 23049;
   hmiStns[1].wip[6].pnCode[0] := 0;
   hmiStns[1].wip[6].pnCode[1] := 243000;
   hmiStns[1].wip[6].pnCode[2] := 70000;
   hmiStns[1].wip[6].pnCode[3] := 73000;
   hmiStns[1].wip[6].pnCode[4] := 0;
   hmiStns[1].wip[6].pnCode[5] := 58000;
   hmiStns[1].wip[6].pnCode[6] := 41000;
   hmiStns[1].wip[6].pnCode[7] := 72000;
   hmiStns[1].wip[7].wipCode := 75057;
   hmiStns[1].wip[7].pnCode[0] := 0;
   hmiStns[1].wip[7].pnCode[1] := 243000;
   hmiStns[1].wip[7].pnCode[2] := 228000;
   hmiStns[1].wip[7].pnCode[3] := 231000;
   hmiStns[1].wip[7].pnCode[4] := 0;
   hmiStns[1].wip[7].pnCode[5] := 229000;
   hmiStns[1].wip[7].pnCode[6] := 227000;
   hmiStns[1].wip[7].pnCode[7] := 230000;
   hmiStns[1].wip[8].wipCode := 76058;
   hmiStns[1].wip[8].pnCode[0] := 0;
   hmiStns[1].wip[8].pnCode[1] := 243000;
   hmiStns[1].wip[8].pnCode[2] := 233000;
   hmiStns[1].wip[8].pnCode[3] := 0;
   hmiStns[1].wip[8].pnCode[4] := 0;
   hmiStns[1].wip[8].pnCode[5] := 229000;
   hmiStns[1].wip[8].pnCode[6] := 232000;
   hmiStns[1].wip[8].pnCode[7] := 231000;
   hmiStns[1].wip[9].wipCode := 77055;
   hmiStns[1].wip[9].pnCode[0] := 0;
   hmiStns[1].wip[9].pnCode[1] := 243000;
   hmiStns[1].wip[9].pnCode[2] := 236000;
   hmiStns[1].wip[9].pnCode[3] := 0;
   hmiStns[1].wip[9].pnCode[4] := 0;
   hmiStns[1].wip[9].pnCode[5] := 237000;
   hmiStns[1].wip[9].pnCode[6] := 234000;
   hmiStns[1].wip[9].pnCode[7] := 235000;
   hmiStns[1].wip[10].wipCode := 78055;
   hmiStns[1].wip[10].pnCode[0] := 0;
   hmiStns[1].wip[10].pnCode[1] := 243000;
   hmiStns[1].wip[10].pnCode[2] := 164000;
   hmiStns[1].wip[10].pnCode[3] := 0;
   hmiStns[1].wip[10].pnCode[4] := 0;
   hmiStns[1].wip[10].pnCode[5] := 165000;
   hmiStns[1].wip[10].pnCode[6] := 234000;
   hmiStns[1].wip[10].pnCode[7] := 235000;
   hmiStns[1].wip[11].wipCode := 79048;
   hmiStns[1].wip[11].pnCode[0] := 0;
   hmiStns[1].wip[11].pnCode[1] := 243000;
   hmiStns[1].wip[11].pnCode[2] := 201000;
   hmiStns[1].wip[11].pnCode[3] := 0;
   hmiStns[1].wip[11].pnCode[4] := 0;
   hmiStns[1].wip[11].pnCode[5] := 200000;
   hmiStns[1].wip[11].pnCode[6] := 234000;
   hmiStns[1].wip[11].pnCode[7] := 235000;
   hmiStns[1].wip[12].wipCode := 80054;
   hmiStns[1].wip[12].pnCode[0] := 0;
   hmiStns[1].wip[12].pnCode[1] := 243000;
   hmiStns[1].wip[12].pnCode[2] := 240000;
   hmiStns[1].wip[12].pnCode[3] := 0;
   hmiStns[1].wip[12].pnCode[4] := 0;
   hmiStns[1].wip[12].pnCode[5] := 241000;
   hmiStns[1].wip[12].pnCode[6] := 238000;
   hmiStns[1].wip[12].pnCode[7] := 239000;
   hmiStns[1].wip[13].wipCode := 20050;
   hmiStns[1].wip[13].pnCode[0] := 0;
   hmiStns[1].wip[13].pnCode[1] := 243000;
   hmiStns[1].wip[13].pnCode[2] := 70000;
   hmiStns[1].wip[13].pnCode[3] := 72000;
   hmiStns[1].wip[13].pnCode[4] := 0;